   
   IF Sbr_IN_xHeadPos THEN
   	Z300_BufferPlate.rgtPlate[Sbr_IN_dCapIndex].tData.tFlag.tConveyor.xDoneHeadPositioning := 1;
   	IF (Z300_BufferPlate.rgtPlate[Sbr_IN_dCapIndex].tData.dTotalCaps > 1) AND (Z300_BufferPlate.rgtPlate[Sbr_IN_dCapIndex].tTracking.dNextCapIndex > 0) THEN
   		JSR(sbrTrackingPositioningDone,2,Z300_BufferPlate.rgtPlate[Sbr_IN_dCapIndex].tTracking.dNextCapIndex,Sbr_IN_xHeadPos);
   	END_IF;
   ELSE
   	Z300_BufferPlate.rgtPlate[Sbr_IN_dCapIndex].tData.tFlag.tConveyor.xDoneTailPositioning := 1;
   	IF (Z300_BufferPlate.rgtPlate[Sbr_IN_dCapIndex].tData.dTotalCaps > 1) AND (Z300_BufferPlate.rgtPlate[Sbr_IN_dCapIndex].tTracking.dNextCapIndex > 0) THEN
   		JSR(sbrTrackingPositioningDone,2,Z300_BufferPlate.rgtPlate[Sbr_IN_dCapIndex].tTracking.dNextCapIndex,Sbr_IN_xHeadPos);
   	END_IF;
   END_IF;
   
   /*
   Z300_BufferPlate.rgtPlate[Sbr_IN_dCapIndex].tTracking.dPosition_cmm := Sbr_IN_Position - Z300_BufferPlate.rgtPlate[Sbr_IN_dCapIndex].tTracking.dLength_cmm / 2;
   ///////////////// CONVOY SYNCHRONIZATION
   IF (Z300_BufferPlate.rgtPlate[Sbr_IN_dCapIndex].tData.dTotalCaps > 1) AND (Z300_BufferPlate.rgtPlate[Sbr_IN_dCapIndex].tData.dCapIndex = 0) THEN
   	JSR(sbrZ300ConvoySynchronization,1,Sbr_IN_dCapIndex);
   END_IF;
   */
   
END_ROUTINE

ROUTINE sbrTrackingPositioningStart   (* structured text *)
   
   SBR(Sbr_IN_dCapIndex,Sbr_IN_xHeadPos);
   
   IF Sbr_IN_xHeadPos THEN
   	Z300_BufferPlate.rgtPlate[Sbr_IN_dCapIndex].tData.tFlag.tConveyor.xDoneHeadPositioning := 0;
   	IF (Z300_BufferPlate.rgtPlate[Sbr_IN_dCapIndex].tData.dTotalCaps > 1) AND (Z300_BufferPlate.rgtPlate[Sbr_IN_dCapIndex].tTracking.dNextCapIndex > 0) THEN
   		JSR(sbrTrackingPositioningDone,2,Z300_BufferPlate.rgtPlate[Sbr_IN_dCapIndex].tTracking.dNextCapIndex,Sbr_IN_xHeadPos);
   	END_IF;
   ELSE
   	Z300_BufferPlate.rgtPlate[Sbr_IN_dCapIndex].tData.tFlag.tConveyor.xDoneTailPositioning := 0;
   	IF (Z300_BufferPlate.rgtPlate[Sbr_IN_dCapIndex].tData.dTotalCaps > 1) AND (Z300_BufferPlate.rgtPlate[Sbr_IN_dCapIndex].tTracking.dNextCapIndex > 0) THEN
   		JSR(sbrTrackingPositioningDone,2,Z300_BufferPlate.rgtPlate[Sbr_IN_dCapIndex].tTracking.dNextCapIndex,Sbr_IN_xHeadPos);
   	END_IF;
   END_IF;
   
END_ROUTINE

ROUTINE sbrTrackingShift   (* structured text *)
   
   FOR TMP_dIndexCap:=0 TO CONST_tPlant.dMaxNumPlates - 1 DO
   	TMP_xTailFound := 0;
   	TMP_xCenterFound := 0;
   	TMP_OUT_xPlateEndTracking := 0;
   	SIZE(Z300_LineTracking.rgtTrkConv[0],0,TMP_dLineSize);
   
   	//Check Tracking Data Present
   	IF (Z300_BufferPlate.rgtPlate[TMP_dIndexCap].tTracking.dPosition_cmm < Z300_dEndTrackingPosition) AND (Z300_BufferPlate.rgtPlate[TMP_dIndexCap].tTracking.dLength_cmm > 0) THEN
   	    TMP_dStepAdvMotor := Z300_BufferPlate.rgtPlate[TMP_dIndexCap].tTracking.dIndexMotorStepAdv;
   		IF NOT Z300_BufferPlate.rgtPlate[TMP_dIndexCap].tTracking.xNotConsConvTrk THEN
   			IF Z300_BufferPlate.rgtPlate[TMP_dIndexCap].tTracking.dLastConv > 0 THEN
   		        TMP_dLastConv := Z300_BufferPlate.rgtPlate[TMP_dIndexCap].tTracking.dLastConv;
   		        Z300_BufferPlate.rgtPlate[TMP_dIndexCap].tTracking.dLastConv := 0;
   
   		        FOR TMP_dIndexConv := TMP_dLastConv - 1 TO TMP_dLastConv + 1 DO
   		            IF (Z300_BufferPlate.rgtPlate[TMP_dIndexCap].tTracking.dPosition_cmm >= Z300_LineTracking.rgtTrkConv[TMP_dIndexConv].dStartPosition_cmm
   						OR (Z300_BufferPlate.rgtPlate[TMP_dIndexCap].tTracking.dPosition_cmm <= Z300_LineTracking.rgtTrkConv[TMP_dIndexConv].dStartPosition_cmm AND TMP_dIndexConv = 0 ))
   		                   AND Z300_BufferPlate.rgtPlate[TMP_dIndexCap].tTracking.dPosition_cmm <= Z300_LineTracking.rgtTrkConv[TMP_dIndexConv].dEndPosition_cmm THEN
   		                IF NOT Z300_BufferPlate.rgtPlate[TMP_dIndexCap].tTracking.xHoldAdvancement THEN
   							IF Z300_Conveyor_Conf[TMP_dIndexConv].dMotorNumber > 0 THEN
   								TMP_dStepAdvMotor := Z300_BufferPlate.rgtPlate[TMP_dIndexCap].tTracking.dIndexMotorStepAdv;
   							ELSE //One motor presence considerate the plate on the first
   								TMP_dStepAdvMotor := 0;
   							END_IF;
   		                    Z300_BufferPlate.rgtPlate[TMP_dIndexCap].tTracking.dPosition_cmm := Z300_BufferPlate.rgtPlate[TMP_dIndexCap].tTracking.dPosition_cmm + Z300_LineTracking.rgtTrkConv[TMP_dIndexConv].dStepAdv_cmm[TMP_dStepAdvMotor];
   		                END_IF;
   		                Z300_BufferPlate.rgtPlate[TMP_dIndexCap].tTracking.dLastConv := TMP_dIndexConv;
   		                EXIT;
   		            END_IF;
   		        END_FOR;
   
   		     // Global Search
   		     ELSE
   		         FOR TMP_dIndexConv := 0 TO TMP_dLineSize - 1 DO
   		             IF (Z300_BufferPlate.rgtPlate[TMP_dIndexCap].tTracking.dPosition_cmm >= Z300_LineTracking.rgtTrkConv[TMP_dIndexConv].dStartPosition_cmm OR
   		                 (Z300_BufferPlate.rgtPlate[TMP_dIndexCap].tTracking.dPosition_cmm <= Z300_LineTracking.rgtTrkConv[TMP_dIndexConv].dStartPosition_cmm AND TMP_dIndexConv = 0 ))
   		                 AND Z300_BufferPlate.rgtPlate[TMP_dIndexCap].tTracking.dPosition_cmm <= Z300_LineTracking.rgtTrkConv[TMP_dIndexConv].dEndPosition_cmm THEN
   		                IF NOT Z300_BufferPlate.rgtPlate[TMP_dIndexCap].tTracking.xHoldAdvancement THEN
   							IF Z300_Conveyor_Conf[TMP_dIndexConv].dMotorNumber > 0 THEN
   								TMP_dStepAdvMotor := Z300_BufferPlate.rgtPlate[TMP_dIndexCap].tTracking.dIndexMotorStepAdv;
   							ELSE //One motor presence considerate the plate on the first
   								TMP_dStepAdvMotor := 0;
   							END_IF;
   		                    Z300_BufferPlate.rgtPlate[TMP_dIndexCap].tTracking.dPosition_cmm := Z300_BufferPlate.rgtPlate[TMP_dIndexCap].tTracking.dPosition_cmm + Z300_LineTracking.rgtTrkConv[TMP_dIndexConv].dStepAdv_cmm[TMP_dStepAdvMotor];
   		                END_IF;
   		                Z300_BufferPlate.rgtPlate[TMP_dIndexCap].tTracking.dLastConv := TMP_dIndexConv;
   		                EXIT;
   		            END_IF;
   		        END_FOR;
   		    END_IF;
   	    ELSE
   			IF NOT Z300_BufferPlate.rgtPlate[TMP_dIndexCap].tTracking.xHoldAdvancement THEN
               	TMP_dIndexConv := Z300_BufferPlate.rgtPlate[TMP_dIndexCap].tTracking.dIndexConvNotCons;
               	IF Z300_Conveyor_Conf[TMP_dIndexConv].dMotorNumber > 0 THEN
   					TMP_dStepAdvMotor := Z300_BufferPlate.rgtPlate[TMP_dIndexCap].tTracking.dIndexMotorStepAdv;
   				ELSE //One motor presence considerate the plate on the first
   					TMP_dStepAdvMotor := 0;
   				END_IF;
               	Z300_BufferPlate.rgtPlate[TMP_dIndexCap].tTracking.dPosition_cmm := Z300_BufferPlate.rgtPlate[TMP_dIndexCap].tTracking.dPosition_cmm + Z300_LineTracking.rgtTrkConv[TMP_dIndexConv].dStepAdv_cmm[TMP_dStepAdvMotor];
           	END_IF;
           	Z300_BufferPlate.rgtPlate[TMP_dIndexCap].tTracking.dLastConv := TMP_dIndexConv;
   		END_IF;
   
   	    TMP_dLastConvTail := Z300_BufferPlate.rgtPlate[TMP_dIndexCap].tTracking.dLastConvTail;
   	    Z300_BufferPlate.rgtPlate[TMP_dIndexCap].tTracking.dLastConvTail := 0;
   	    TMP_xTailFound := 0;
   	    TMP_xCenterFound := 0;
   	    FOR TMP_dIndexConv := TMP_dLastConvTail TO TMP_dLineSize - 1 DO
   
               TMP_dIndexCapConv := Z300_LineTracking.rgtTrkConv[TMP_dIndexConv].dIndexCaps;// - 1;
   
   			IF TMP_dIndexCapConv < CONST_tPlant.dNumCapsConveyor THEN
   	            TMP_dPosTail_cmm := Z300_BufferPlate.rgtPlate[TMP_dIndexCap].tTracking.dPosition_cmm - (Z300_BufferPlate.rgtPlate[TMP_dIndexCap].tTracking.dLength_cmm / 2);
   	            TMP_dPosHead_cmm := Z300_BufferPlate.rgtPlate[TMP_dIndexCap].tTracking.dPosition_cmm + (Z300_BufferPlate.rgtPlate[TMP_dIndexCap].tTracking.dLength_cmm/ 2);
   	            TMP_dPos_cmm := Z300_BufferPlate.rgtPlate[TMP_dIndexCap].tTracking.dPosition_cmm - (Z300_BufferPlate.rgtPlate[TMP_dIndexCap].tTracking.dLength_cmm / 2);
   
   	            //Tail
   	            IF TMP_dPos_cmm >= Z300_LineTracking.rgtTrkConv[TMP_dIndexConv].dStartPosition_cmm
   					AND TMP_dPos_cmm < Z300_LineTracking.rgtTrkConv[TMP_dIndexConv].dEndPosition_cmm  AND NOT TMP_xTailFound THEN
   	                IF TMP_dPos_cmm >= 0 AND TMP_dPos_cmm < Z300_dEndTrackingPosition THEN
   	                    Z300_LineTracking.rgtTrkConv[TMP_dIndexConv].Cap[TMP_dIndexCapConv].xTail := 1;
   	                    Z300_LineTracking.rgtTrkConv[TMP_dIndexConv].Cap[TMP_dIndexCapConv].xPresence := 1;
   	                    Z300_LineTracking.rgtTrkConv[TMP_dIndexConv].Cap[TMP_dIndexCapConv].dTailPos_cmm := TMP_dPos_cmm;
   	                    Z300_LineTracking.rgtTrkConv[TMP_dIndexConv].Cap[TMP_dIndexCapConv].dTailPosConv_cmm := TMP_dPos_cmm - Z300_LineTracking.rgtTrkConv[TMP_dIndexConv].dStartPosition_cmm;
   	                    Z300_LineTracking.rgtTrkConv[TMP_dIndexConv].Cap[TMP_dIndexCapConv].dPointer := TMP_dIndexCap;
   	                    Z300_LineTracking.rgtTrkConv[TMP_dIndexConv].Cap[TMP_dIndexCapConv].dPresenceHead_cmm := TMP_dPosHead_cmm;
   	                    Z300_LineTracking.rgtTrkConv[TMP_dIndexConv].Cap[TMP_dIndexCapConv].dPresenceTail_cmm := TMP_dPosTail_cmm;
   	                    Z300_BufferPlate.rgtPlate[TMP_dIndexCap].tTracking.dIndexConvTail := TMP_dIndexConv;
   	                    TMP_xTailFound := 1;
   	                    Z300_BufferPlate.rgtPlate[TMP_dIndexCap].tTracking.dLastConvTail := TMP_dIndexConv;
   	                    Z300_BufferPlate.rgtPlate[TMP_dIndexCap].tTracking.dIndexCapInConvTail := TMP_dIndexCap;
   	                    Z300_BufferPlate.rgtPlate[TMP_dIndexCap].tTracking.dPositionTail_cmm := TMP_dPos_cmm;
   	                END_IF;
   	            END_IF;
   
   	            // Center Position
   	            TMP_dPosTail_cmm := Z300_BufferPlate.rgtPlate[TMP_dIndexCap].tTracking.dPosition_cmm - (Z300_BufferPlate.rgtPlate[TMP_dIndexCap].tTracking.dLength_cmm / 2);
   	            TMP_dPosHead_cmm := Z300_BufferPlate.rgtPlate[TMP_dIndexCap].tTracking.dPosition_cmm + (Z300_BufferPlate.rgtPlate[TMP_dIndexCap].tTracking.dLength_cmm / 2);
   	            TMP_dPos_cmm := Z300_BufferPlate.rgtPlate[TMP_dIndexCap].tTracking.dPosition_cmm;
   	            IF TMP_dPos_cmm >= Z300_LineTracking.rgtTrkConv[TMP_dIndexConv].dStartPosition_cmm
   					AND TMP_dPos_cmm < Z300_LineTracking.rgtTrkConv[TMP_dIndexConv].dEndPosition_cmm AND NOT TMP_xCenterFound THEN
   	                IF TMP_dPos_cmm >= Z300_dStartTrackingPosition AND TMP_dPos_cmm < Z300_dEndTrackingPosition THEN
   	                    Z300_LineTracking.rgtTrkConv[TMP_dIndexConv].Cap[TMP_dIndexCapConv].xCenter := 1;
   	                    Z300_LineTracking.rgtTrkConv[TMP_dIndexConv].Cap[TMP_dIndexCapConv].xPresence := 1;
   	                    Z300_LineTracking.rgtTrkConv[TMP_dIndexConv].Cap[TMP_dIndexCapConv].dCenterPos_cmm := TMP_dPos_cmm;
   	                    Z300_LineTracking.rgtTrkConv[TMP_dIndexConv].Cap[TMP_dIndexCapConv].dCenterPosConv_cmm := TMP_dPos_cmm - Z300_LineTracking.rgtTrkConv[TMP_dIndexConv].dStartPosition_cmm;
   	                    Z300_LineTracking.rgtTrkConv[TMP_dIndexConv].Cap[TMP_dIndexCapConv].dPointer := TMP_dIndexCap;
   	                    Z300_LineTracking.rgtTrkConv[TMP_dIndexConv].Cap[TMP_dIndexCapConv].dPresenceHead_cmm := TMP_dPosHead_cmm;
   	                    Z300_LineTracking.rgtTrkConv[TMP_dIndexConv].Cap[TMP_dIndexCapConv].dPresenceTail_cmm := TMP_dPosTail_cmm;
   	                    TMP_xCenterFound := 1;
   	                END_IF;
   	            END_IF;
   
   	            //Plate Presence
   	            TMP_dPosTail_cmm := Z300_BufferPlate.rgtPlate[TMP_dIndexCap].tTracking.dPosition_cmm - (Z300_BufferPlate.rgtPlate[TMP_dIndexCap].tTracking.dLength_cmm / 2);
   	            TMP_dPosHead_cmm := Z300_BufferPlate.rgtPlate[TMP_dIndexCap].tTracking.dPosition_cmm + (Z300_BufferPlate.rgtPlate[TMP_dIndexCap].tTracking.dLength_cmm / 2);
   	            IF TMP_dPosTail_cmm <= Z300_LineTracking.rgtTrkConv[TMP_dIndexConv].dStartPosition_cmm
   					AND TMP_dPosHead_cmm >= Z300_LineTracking.rgtTrkConv[TMP_dIndexConv].dEndPosition_cmm  THEN
   	                IF TMP_dPos_cmm >= Z300_dStartTrackingPosition AND TMP_dPos_cmm < Z300_dEndTrackingPosition THEN
   	                    Z300_LineTracking.rgtTrkConv[TMP_dIndexConv].Cap[TMP_dIndexCapConv].xPresence := 1;
   	                    Z300_LineTracking.rgtTrkConv[TMP_dIndexConv].Cap[TMP_dIndexCapConv].dCenterPos_cmm := TMP_dPos_cmm;
   	                    Z300_LineTracking.rgtTrkConv[TMP_dIndexConv].Cap[TMP_dIndexCapConv].dPresenceHead_cmm := TMP_dPosHead_cmm;
   	                    Z300_LineTracking.rgtTrkConv[TMP_dIndexConv].Cap[TMP_dIndexCapConv].dPresenceTail_cmm := TMP_dPosTail_cmm;
   	                    Z300_LineTracking.rgtTrkConv[TMP_dIndexConv].Cap[TMP_dIndexCapConv].dCenterPosConv_cmm := TMP_dPos_cmm - Z300_LineTracking.rgtTrkConv[TMP_dIndexConv].dStartPosition_cmm;
   	                    Z300_LineTracking.rgtTrkConv[TMP_dIndexConv].Cap[TMP_dIndexCapConv].dPointer := TMP_dIndexCap;
   	                    TMP_xPlateFound := 1;
   	                END_IF;
   	            END_IF;
   
   	            // Head Position
   	            TMP_dPosTail_cmm := Z300_BufferPlate.rgtPlate[TMP_dIndexCap].tTracking.dPosition_cmm - (Z300_BufferPlate.rgtPlate[TMP_dIndexCap].tTracking.dLength_cmm / 2);
   	            TMP_dPosHead_cmm := Z300_BufferPlate.rgtPlate[TMP_dIndexCap].tTracking.dPosition_cmm + (Z300_BufferPlate.rgtPlate[TMP_dIndexCap].tTracking.dLength_cmm / 2);
   	            TMP_dPos_cmm := Z300_BufferPlate.rgtPlate[TMP_dIndexCap].tTracking.dPosition_cmm + (Z300_BufferPlate.rgtPlate[TMP_dIndexCap].tTracking.dLength_cmm / 2);
   	            IF (TMP_dPos_cmm >= Z300_LineTracking.rgtTrkConv[TMP_dIndexConv].dStartPosition_cmm)
   					AND (TMP_dPos_cmm < Z300_LineTracking.rgtTrkConv[TMP_dIndexConv].dEndPosition_cmm) AND TMP_xCenterFound THEN
   	                IF TMP_dPos_cmm >= Z300_dStartTrackingPosition AND TMP_dPos_cmm < Z300_dEndTrackingPosition THEN
   	                    Z300_LineTracking.rgtTrkConv[TMP_dIndexConv].Cap[TMP_dIndexCapConv].xHead := 1;
   	                    Z300_LineTracking.rgtTrkConv[TMP_dIndexConv].Cap[TMP_dIndexCapConv].xPresence := 1;
   	                    Z300_LineTracking.rgtTrkConv[TMP_dIndexConv].Cap[TMP_dIndexCapConv].dHeadPos_cmm := TMP_dPos_cmm;
   	                    Z300_LineTracking.rgtTrkConv[TMP_dIndexConv].Cap[TMP_dIndexCapConv].dHeadPosConv_cmm := TMP_dPos_cmm - Z300_LineTracking.rgtTrkConv[TMP_dIndexConv].dStartPosition_cmm;
   	                    Z300_LineTracking.rgtTrkConv[TMP_dIndexConv].Cap[TMP_dIndexCapConv].dPointer := TMP_dIndexCap;
   	                    Z300_LineTracking.rgtTrkConv[TMP_dIndexConv].Cap[TMP_dIndexCapConv].dPresenceHead_cmm := TMP_dPosHead_cmm;
   	                    Z300_LineTracking.rgtTrkConv[TMP_dIndexConv].Cap[TMP_dIndexCapConv].dPresenceTail_cmm := TMP_dPosTail_cmm;
   	                    //Increment Index Single Caps in the conveyor
   	                    Z300_LineTracking.rgtTrkConv[TMP_dIndexConv].dIndexCaps := Z300_LineTracking.rgtTrkConv[TMP_dIndexConv].dIndexCaps + 1;
   	                    IF Z300_LineTracking.rgtTrkConv[TMP_dIndexConv].dIndexCaps >= CONST_tPlant.dNumCapsConveyor THEN
   	                        Z300_LineTracking.rgtTrkConv[TMP_dIndexConv].dIndexCaps := CONST_tPlant.dNumCapsConveyor - 1;
   	                    END_IF;
   	                    Z300_BufferPlate.rgtPlate[TMP_dIndexCap].tTracking.dIndexConvHead := TMP_dIndexConv;
   	                    Z300_BufferPlate.rgtPlate[TMP_dIndexCap].tTracking.dIndexCapInConvHead := TMP_dIndexCap;
   	                    Z300_BufferPlate.rgtPlate[TMP_dIndexCap].tTracking.dPositionHead_cmm := TMP_dPos_cmm;
   	                    EXIT;
   	                END_IF;
   	            END_IF;
   
   			END_IF;
   
               IF  TMP_xTailFound OR TMP_xCenterFound OR TMP_xPlateFound THEN
                   //Increment Index Single Caps in the conveyor
                   Z300_LineTracking.rgtTrkConv[TMP_dIndexConv].dIndexCaps := Z300_LineTracking.rgtTrkConv[TMP_dIndexConv].dIndexCaps + 1;
                   IF Z300_LineTracking.rgtTrkConv[TMP_dIndexConv].dIndexCaps >= CONST_tPlant.dNumCapsConveyor THEN
                       Z300_LineTracking.rgtTrkConv[TMP_dIndexConv].dIndexCaps := CONST_tPlant.dNumCapsConveyor - 1;
                   END_IF;
               END_IF;
           END_FOR;
       ELSE
   		//plate not more in tracking area
   		TMP_OUT_xPlateEndTracking := Z300_BufferPlate.rgtPlate[TMP_dIndexCap].tTracking.dPosition_cmm >= Z300_dEndTrackingPosition;
   	END_IF;
   
       //write the Output
       Z300_BufferPlate.rgtPlate[TMP_dIndexCap].tTracking.dPosition_cmm := Z300_BufferPlate.rgtPlate[TMP_dIndexCap].tTracking.dPosition_cmm;
   
   	//if plate at end of tracking delete from tracking
   	IF TMP_OUT_xPlateEndTracking THEN
   		COP(AUX_tBufferPlate_NULL,Z300_BufferPlate.rgtPlate[TMP_dIndexCap],1);
   	END_IF;
   END_FOR;
   
END_ROUTINE

ROUTINE sbrTrimWheelTrPositionOppOpSide   (* ladder *)
   0: NOP();
   1: [XIC(M30xTrimWheel[TMP_dIndex].OS_xStartPositioningOppOpSide) ,XIC(M30xTrimWheel[TMP_dIndex].OS_xReqUpdateTargetTranslationOppOpSide) ]ADD(M30xTrimWheel[TMP_dIndex].AUX_dReqTargetPosTranslation_cmm[1],M30xTrimWheel[TMP_dIndex].AUX_dOffsetSingle_cmm[1],M30xTrimWheel[TMP_dIndex].AUX_dFinalTarget_cmm[1]);
   2: GP_PosWindow(GP_PosWindow,M30xTrimWheel[TMP_dIndex].AUX_dFinalTarget_cmm[1],M30xTrimWheel[TMP_dIndex].AUX_dActTransPosition_cmm[1],M30xTrimWheel[TMP_dIndex].CONF_dTolerance_cmm[1],0,M30xTrimWheel[TMP_dIndex].ST_xInPositionOppOpSide);
   3: GP_PosWindow(GP_PosWindow,M30xTrimWheel[TMP_dIndex].AUX_dFinalTarget_cmm[1],M30xTrimWheel[TMP_dIndex].AUX_dActTransPosition_cmm[1],M30xTrimWheel[TMP_dIndex].CONF_dStopCamPos_cmm[1],0,M30xTrimWheel[TMP_dIndex].ST_xInStopCamPositionOppOpSide);
   4: GP_PosWindow(GP_PosWindow,M30xTrimWheel_HMW[TMP_dIndex].rgdPositionManCmd_cmm[1],M30xTrimWheel[TMP_dIndex].AUX_dActTransPosition_cmm[1],M30xTrimWheel[TMP_dIndex].CONF_dSlowDownPos_cmm[1],0,M30xTrimWheel[TMP_dIndex].ST_xInSlowDownManualPosOppOpSide);
   5: GP_PosWindow(GP_PosWindow,M30xTrimWheel_HMW[TMP_dIndex].rgdPositionManCmd_cmm[1],M30xTrimWheel[TMP_dIndex].AUX_dActTransPosition_cmm[1],M30xTrimWheel[TMP_dIndex].CONF_dStopCamPos_cmm[1],0,M30xTrimWheel[TMP_dIndex].ST_xInStopCamManualPositionOppOpSide);
   6: XIC(M30xTrimWheel_HMW[TMP_dIndex].rgxMan.x12)MOV(M30xTrimWheel[TMP_dIndex].CONF_dTrimWheelMaxRange_cmm[1],TMP_dManualTargetPos);
   7: XIC(M30xTrimWheel_HMW[TMP_dIndex].rgxMan.x13)MOV(M30xTrimWheel[TMP_dIndex].CONF_dTrimWheelMinRange_cmm[1],TMP_dManualTargetPos);
   8: GP_PosWindow(GP_PosWindow,TMP_dManualTargetPos,M30xTrimWheel[TMP_dIndex].AUX_dActTransPosition_cmm[1],M30xTrimWheel[TMP_dIndex].CONF_dSlowDownPos_cmm[1],0,M30xTrimWheel[TMP_dIndex].ST_xInSlowDownManualOppOpSide);
   9: GP_PosWindow(GP_PosWindow,TMP_dManualTargetPos,M30xTrimWheel[TMP_dIndex].AUX_dActTransPosition_cmm[1],M30xTrimWheel[TMP_dIndex].CONF_dStopCamPos_cmm[1],0,M30xTrimWheel[TMP_dIndex].ST_xInStopCamManualOppOpSide);
END_ROUTINE

ROUTINE sbrTrimWheelTrPositionOpSide   (* ladder *)
   0: NOP();
   1: [XIC(M30xTrimWheel[TMP_dIndex].OS_xStartPositioningOpSide) ,XIC(M30xTrimWheel[TMP_dIndex].OS_xReqUpdateTargetTranslationOpSide) ]ADD(M30xTrimWheel[TMP_dIndex].AUX_dReqTargetPosTranslation_cmm[0],M30xTrimWheel[TMP_dIndex].AUX_dOffsetSingle_cmm[0],M30xTrimWheel[TMP_dIndex].AUX_dFinalTarget_cmm[0]);
   2: GP_PosWindow(GP_PosWindow,M30xTrimWheel[TMP_dIndex].AUX_dFinalTarget_cmm[0],M30xTrimWheel[TMP_dIndex].AUX_dActTransPosition_cmm[0],M30xTrimWheel[TMP_dIndex].CONF_dTolerance_cmm[0],0,M30xTrimWheel[TMP_dIndex].ST_xInPositionOpSide);
   3: GP_PosWindow(GP_PosWindow,M30xTrimWheel[TMP_dIndex].AUX_dFinalTarget_cmm[0],M30xTrimWheel[TMP_dIndex].AUX_dActTransPosition_cmm[0],M30xTrimWheel[TMP_dIndex].CONF_dStopCamPos_cmm[0],0,M30xTrimWheel[TMP_dIndex].ST_xInStopCamPositionOpSide);
   4: GP_PosWindow(GP_PosWindow,M30xTrimWheel_HMW[TMP_dIndex].rgdPositionManCmd_cmm[0],M30xTrimWheel[TMP_dIndex].AUX_dActTransPosition_cmm[0],M30xTrimWheel[TMP_dIndex].CONF_dSlowDownPos_cmm[0],0,M30xTrimWheel[TMP_dIndex].ST_xInSlowDownManualPosOpSide);
   5: GP_PosWindow(GP_PosWindow,M30xTrimWheel_HMW[TMP_dIndex].rgdPositionManCmd_cmm[0],M30xTrimWheel[TMP_dIndex].AUX_dActTransPosition_cmm[0],M30xTrimWheel[TMP_dIndex].CONF_dStopCamPos_cmm[0],0,M30xTrimWheel[TMP_dIndex].ST_xInStopCamManualPositionOpSide);
   6: XIC(M30xTrimWheel_HMW[TMP_dIndex].rgxMan.x2)MOV(M30xTrimWheel[TMP_dIndex].CONF_dTrimWheelMaxRange_cmm[0],TMP_dManualTargetPos);
   7: XIC(M30xTrimWheel_HMW[TMP_dIndex].rgxMan.x3)MOV(M30xTrimWheel[TMP_dIndex].CONF_dTrimWheelMinRange_cmm[0],TMP_dManualTargetPos);
   8: GP_PosWindow(GP_PosWindow,TMP_dManualTargetPos,M30xTrimWheel[TMP_dIndex].AUX_dActTransPosition_cmm[0],M30xTrimWheel[TMP_dIndex].CONF_dSlowDownPos_cmm[0],0,M30xTrimWheel[TMP_dIndex].ST_xInSlowDownManualOpSide);
   9: GP_PosWindow(GP_PosWindow,TMP_dManualTargetPos,M30xTrimWheel[TMP_dIndex].AUX_dActTransPosition_cmm[0],M30xTrimWheel[TMP_dIndex].CONF_dStopCamPos_cmm[0],0,M30xTrimWheel[TMP_dIndex].ST_xInStopCamManualOpSide);
END_ROUTINE

ROUTINE sbrUpdateTrackingConvoyPosition   (* structured text *)
   SBR(Sbr_IN_dIndexHead,Sbr_IN_Position);
   
   Z300_BufferPlate.rgtPlate[Sbr_IN_dIndexHead].tTracking.dPosition_cmm := Sbr_IN_Position - Z300_BufferPlate.rgtPlate[Sbr_IN_dIndexHead].tTracking.dLength_cmm / 2;
   ///////////////// CONVOY SYNCHRONIZATION
   IF (Z300_BufferPlate.rgtPlate[Sbr_IN_dIndexHead].tData.dTotalCaps > 1) AND (Z300_BufferPlate.rgtPlate[Sbr_IN_dIndexHead].tData.dCapIndex = 0) THEN
   //Search for single caps within the same convoy
   	// Synchronize convoy
   	JSR(sbrZ300ConvoySynchronization,1,Sbr_IN_dIndexHead);
   END_IF;
   
END_ROUTINE

ROUTINE sbrZ300ConvoySynchronization   (* structured text *)
   /*
   //Initialize
   TMP_dPnt1 := Z300_Photocell[TMP_dIndex].tSearchPlate.rgdHeadPointer[0];
   TMP_dPnt2 := Z300_Photocell[TMP_dIndex].tSearchPlate.rgdHeadPointer[1];
   TMP_dPnt3 := Z300_Photocell[TMP_dIndex].tSearchPlate.rgdHeadPointer[2];
   TMP_dPnt4 := Z300_Photocell[TMP_dIndex].tSearchPlate.rgdHeadPointer[3];
   //If convoy in progress synchronize second cap
   IF (Z300_Photocell[TMP_dIndex].tSearchPlate.rgxHead > 1) AND (Z300_BufferPlate.rgtPlate[TMP_dPnt1].tData.dTotalCaps > 1) AND (Z300_BufferPlate.rgtPlate[TMP_dPnt1].tData.rgtCap[0].dIndex = 0)
   AND (Z300_BufferPlate.rgtPlate[TMP_dPnt2].tData.dTotalCaps > 1) AND (Z300_BufferPlate.rgtPlate[TMP_dPnt2].tData.rgtCap[0].dIndex = 1) THEN
   	//Synchronyze also second cap
   	Z300_BufferPlate.rgtPlate[TMP_dPnt2].tTracking.dPosition_cmm := Z300_BufferPlate.rgtPlate[TMP_dPnt1].tTracking.dPosition_cmm
   	- (Z300_BufferPlate.rgtPlate[TMP_dPnt1].tTracking.dLength_cmm / 2)
   	- Z300_BufferPlate.rgtPlate[TMP_dPnt1].tData.dGapCaps_cmm
   	- (Z300_BufferPlate.rgtPlate[TMP_dPnt2].tTracking.dLength_cmm / 2);
   END_IF;
   //If convoy in progress synchronize third cap
   IF (Z300_Photocell[TMP_dIndex].tSearchPlate.rgxHead > 2) AND (Z300_BufferPlate.rgtPlate[TMP_dPnt2].tData.dTotalCaps > 2) AND (Z300_BufferPlate.rgtPlate[TMP_dPnt2].tData.rgtCap[0].dIndex = 1)
   AND (Z300_BufferPlate.rgtPlate[TMP_dPnt3].tData.dTotalCaps > 2) AND (Z300_BufferPlate.rgtPlate[TMP_dPnt3].tData.rgtCap[0].dIndex = 2) THEN
   	//Synchronyze also third cap
   	Z300_BufferPlate.rgtPlate[TMP_dPnt3].tTracking.dPosition_cmm := Z300_BufferPlate.rgtPlate[TMP_dPnt2].tTracking.dPosition_cmm
   	- (Z300_BufferPlate.rgtPlate[TMP_dPnt2].tTracking.dLength_cmm / 2)
   	- Z300_BufferPlate.rgtPlate[TMP_dPnt2].tData.dGapCaps_cmm
   	- (Z300_BufferPlate.rgtPlate[TMP_dPnt3].tTracking.dLength_cmm / 2);
   END_IF;
   //If convoy in progress synchronize fourth cap
   IF (Z300_Photocell[TMP_dIndex].tSearchPlate.rgxHead > 3) AND (Z300_BufferPlate.rgtPlate[TMP_dPnt3].tData.dTotalCaps > 3) AND (Z300_BufferPlate.rgtPlate[TMP_dPnt3].tData.rgtCap[0].dIndex = 2)
   AND (Z300_BufferPlate.rgtPlate[TMP_dPnt4].tData.dTotalCaps > 3) AND (Z300_BufferPlate.rgtPlate[TMP_dPnt4].tData.rgtCap[0].dIndex = 3) THEN
   	//Synchronyze also fourth cap
   	Z300_BufferPlate.rgtPlate[TMP_dPnt4].tTracking.dPosition_cmm := Z300_BufferPlate.rgtPlate[TMP_dPnt3].tTracking.dPosition_cmm
   	- (Z300_BufferPlate.rgtPlate[TMP_dPnt3].tTracking.dLength_cmm / 2)
   	- Z300_BufferPlate.rgtPlate[TMP_dPnt3].tData.dGapCaps_cmm
   	- (Z300_BufferPlate.rgtPlate[TMP_dPnt4].tTracking.dLength_cmm / 2);
   END_IF;
   */
   
   SBR(Sbr_IN_dCapIndex);
   
   TMP_dNextCap := Z300_BufferPlate.rgtPlate[Sbr_IN_dCapIndex].tTracking.dNextCapIndex;
   IF TMP_dNextCap > 0 THEN
   	Z300_BufferPlate.rgtPlate[TMP_dNextCap].tTracking.dPosition_cmm := Z300_BufferPlate.rgtPlate[Sbr_IN_dCapIndex].tTracking.dPosition_cmm - Z300_BufferPlate.rgtPlate[Sbr_IN_dCapIndex].tTracking.dLength_cmm / 2
   	- Z300_BufferPlate.rgtPlate[Sbr_IN_dCapIndex].tData.dGapCaps_cmm - Z300_BufferPlate.rgtPlate[TMP_dNextCap].tTracking.dLength_cmm / 2;
   	JSR(sbrZ300ConvoySynchronization,1,TMP_dNextCap);
   END_IF;
   
END_ROUTINE

ROUTINE ScadaPlate_Logic   (* structured text *)
   
   TMP_xLastModalityLoadBwd := 0;
   TMP_xLastModalityUnloadBwd := 0;
   TMP_xYWithBarycenter := 1;
   TMP_xYInversionLite := 1;
   
   TMP_dCulletMask := CONST_rgdDestMask[24];
   FOR TMP_dIndexPlate := 0 TO CONST_tPlant.dMaxNumPlates - 1 DO
   	//Write data
   	//Calculate Head Position
   	TMP_dHeadPosition_mm := Z300_BufferPlate.rgtPlate[TMP_dIndexPlate].tTracking.dPositionHead_cmm / 100;
   	TMP_dConveyorLength := Z300_dEndTrackingPosition/ 100;
   	TMP_dWidth_mm := Z300_Conveyor_Conf[0].dWidthConveyor_cmm / 100;
   
   	//Init counter cap (always only one cap on line tracking)
   	TMP_dCap := 0;
   
   	//Init counter lite
   	TMP_dLite := 0;
   
   	FOR TMP_dLite := 0 TO CONST_tPlant.dNumLitesMaxCap - 1 DO
   	    IF Z300_BufferPlate.rgtPlate[TMP_dIndexPlate].tData.rgtCap[TMP_dCap].rgtLite[TMP_dLite].dID <> 0 AND NOT Z300_BufferPlate.rgtPlate[TMP_dIndexPlate].tTracking.xNotShownInScada THEN
   	        TMP_dLiteInv := CONST_tPlant.dNumLitesMaxCap - 1 - TMP_dLite;
   
   	        //Plate
   	        Z300_Scada_Continuous.rgtPlate[TMP_dIndexPlate].rgtCap[TMP_dCap].rgtLite[TMP_dLite].dPlateId := Z300_BufferPlate.rgtPlate[TMP_dIndexPlate].tData.rgtCap[TMP_dCap].rgtLite[TMP_dLite].dID;
   	        //Production ID
   	        Z300_Scada_Continuous.rgtPlate[TMP_dIndexPlate].rgtCap[TMP_dCap].rgtLite[TMP_dLite].dProductionID := Z300_BufferPlate.rgtPlate[TMP_dIndexPlate].tData.rgtCap[TMP_dCap].rgtLite[TMP_dLite].dProductionID;
   	        //Plate lenght
   	        Z300_Scada_Continuous.rgtPlate[TMP_dIndexPlate].rgtCap[TMP_dCap].rgtLite[TMP_dLite].dPlateLength_mm := Z300_BufferPlate.rgtPlate[TMP_dIndexPlate].tData.rgtCap[TMP_dCap].dLength_cmm / 100;
   	        //Plate widht
   	        Z300_Scada_Continuous.rgtPlate[TMP_dIndexPlate].rgtCap[TMP_dCap].rgtLite[TMP_dLite].dPlateWidth_mm := Z300_BufferPlate.rgtPlate[TMP_dIndexPlate].tData.rgtCap[TMP_dCap].rgtLite[TMP_dLite].dWidth_cmm / 100;
   
   	        //Init the value of Destination/Source/Alternative/SecondDestination
   	        TMP_xPresenceDestination := 0;
   	        TMP_xPresenceAlternative := 0;
   	        //TMP_xPresenceSource := 0;
   	        TMP_xPresenceSecondDestination := 0;
   
   	        //Destination
   	        FOR TMP_dCountDest := 0 TO 31 DO
   	            //Main Destination
   	            IF Z300_BufferPlate.rgtPlate[TMP_dIndexPlate].tData.rgtCap[TMP_dCap].rgtLite[TMP_dLite].tDestination.rgxMain.[TMP_dCountDest] THEN
   	                Z300_Scada_Continuous.rgtPlate[TMP_dIndexPlate].rgtCap[TMP_dCap].rgtLite[TMP_dLite].dDestination := TMP_dCountDest + 1;
   	                TMP_xPresenceDestination := 1;
   	            END_IF;
   	            ////Source
   				//IF INO_tPlate.tData.rgtCap[TMP_dCap].rgtLite[TMP_dLite].
   	            //IF INO_tPlate.tData.rgtCap[TMP_dCap].rgtLite[TMP_dLite].tSource.rgxOrigin.[TMP_dCountDest] THEN
   	            //    INO_tScada_Continuous.rgtPlate[IN_dIndexPlate].rgtCap[TMP_dCap].rgtLite[TMP_dLite].dSource := TMP_dCountDest + 1;
   	            //    TMP_xPresenceSource := 1;
   	            //END_IF;
   	            //Alternative Destination
   	            IF Z300_BufferPlate.rgtPlate[TMP_dIndexPlate].tData.rgtCap[TMP_dCap].rgtLite[TMP_dLite].tDestination.rgxAlternative.[TMP_dCountDest] THEN
   	                Z300_Scada_Continuous.rgtPlate[TMP_dIndexPlate].rgtCap[TMP_dCap].rgtLite[TMP_dLite].dAlternative := TMP_dCountDest + 1;
   	                TMP_xPresenceAlternative := 1;
   	            END_IF;
   	            //Second Destination
   	            IF Z300_BufferPlate.rgtPlate[TMP_dIndexPlate].tData.rgtCap[TMP_dCap].rgtLite[TMP_dLite].tDestination.rgxAlternative.[TMP_dCountDest] THEN
   	                Z300_Scada_Continuous.rgtPlate[TMP_dIndexPlate].rgtCap[TMP_dCap].rgtLite[TMP_dLite].dSecondDestination := TMP_dCountDest + 1;
   	                TMP_xPresenceSecondDestination := 1;
   	            END_IF;
   	        END_FOR;
   			//IF Z300_BufferPlate.rgtPlate[TMP_dIndexPlate].tData.rgtCap[TMP_dCap].rgtLite[TMP_dLite].tDestination.rgxMain = CONST_rgdDestMask[24] THEN
   	        //    Z300_Scada_Continuous.rgtPlate[TMP_dIndexPlate].rgtCap[TMP_dCap].rgtLite[TMP_dLite].dDestination := CONST_rgdDestMask[24];
   	        //END_IF;
   	        IF NOT TMP_xPresenceDestination THEN
   	            Z300_Scada_Continuous.rgtPlate[TMP_dIndexPlate].rgtCap[TMP_dCap].rgtLite[TMP_dLite].dDestination := 0;
   	        END_IF;
   	        IF NOT TMP_xPresenceAlternative THEN
   	            Z300_Scada_Continuous.rgtPlate[TMP_dIndexPlate].rgtCap[TMP_dCap].rgtLite[TMP_dLite].dAlternative := 0;
   	        END_IF;
   	        IF NOT TMP_xPresenceSecondDestination THEN
   	            Z300_Scada_Continuous.rgtPlate[TMP_dIndexPlate].rgtCap[TMP_dCap].rgtLite[TMP_dLite].dSecondDestination := 0;
   	        END_IF;
   	        //IF NOT TMP_xPresenceSource THEN
   	            Z300_Scada_Continuous.rgtPlate[TMP_dIndexPlate].rgtCap[TMP_dCap].rgtLite[TMP_dLite].dSource := 0;
   	        //END_IF;
   
   	        ////Set origin to 0 in case of destination is <> 0
   	        //IF INO_tScada_Continuous.rgtPlate[IN_dIndexPlate].rgtCap[TMP_dCap].rgtLite[TMP_dLite].dDestination <> 0 THEN
   	        //    INO_tScada_Continuous.rgtPlate[IN_dIndexPlate].rgtCap[TMP_dCap].rgtLite[TMP_dLite].dSource := 0;
   	        //END_IF;
   
   	        //Position x (Forward)
   	        IF NOT TMP_xLastModalityLoadBwd AND NOT TMP_xLastModalityUnloadBwd THEN
   	            //Tail
   	            Z300_Scada_Continuous.rgtPlate[TMP_dIndexPlate].rgtCap[TMP_dCap].rgtLite[TMP_dLite].dTail_PosX_mm := TMP_dHeadPosition_mm - (Z300_BufferPlate.rgtPlate[TMP_dIndexPlate].tData.rgtCap[TMP_dCap].dLength_cmm / 100);
   
   	            //Head
   	            Z300_Scada_Continuous.rgtPlate[TMP_dIndexPlate].rgtCap[TMP_dCap].rgtLite[TMP_dLite].dHead_PosX_mm := TMP_dHeadPosition_mm;
   	        END_IF;
   
   	        //Position x (Backward)
   	        //Head
   
   	        IF TMP_xLastModalityLoadBwd OR TMP_xLastModalityUnloadBwd THEN
   	            //  Head
   	            Z300_Scada_Continuous.rgtPlate[TMP_dIndexPlate].rgtCap[TMP_dCap].rgtLite[TMP_dLite].dHead_PosX_mm := TMP_dConveyorLength - TMP_dHeadPosition_mm + (Z300_BufferPlate.rgtPlate[TMP_dIndexPlate].tData.dLength_cmm / 100);
   
   	            //  Tail
   	            Z300_Scada_Continuous.rgtPlate[TMP_dIndexPlate].rgtCap[TMP_dCap].rgtLite[TMP_dLite].dTail_PosX_mm :=
   	            Z300_Scada_Continuous.rgtPlate[TMP_dIndexPlate].rgtCap[TMP_dCap].rgtLite[TMP_dLite].dHead_PosX_mm - (Z300_BufferPlate.rgtPlate[TMP_dIndexPlate].tData.rgtCap[TMP_dCap].dLength_cmm / 100);
   	        END_IF;
   
   	        //Position Y
   
   	        //Barycenter not used, without inversion (IN FC)
   	        IF NOT TMP_xYWithBarycenter AND NOT TMP_xYInversionLite THEN
   	            IF TMP_dLite < 1 THEN
   	                Z300_Scada_Continuous.rgtPlate[TMP_dIndexPlate].rgtCap[TMP_dCap].rgtLite[TMP_dLite].dPositionY_mm :=
   	                ((TMP_dWidth_mm / 2) - (Z300_BufferPlate.rgtPlate[TMP_dIndexPlate].tData.rgtCap[TMP_dCap].dWidth_cmm / 100) / 2);
   	            ELSE
   	                Z300_Scada_Continuous.rgtPlate[TMP_dIndexPlate].rgtCap[TMP_dCap].rgtLite[TMP_dLite].dPositionY_mm := Z300_Scada_Continuous.rgtPlate[TMP_dIndexPlate].rgtCap[TMP_dCap].rgtLite[TMP_dLite - 1].dPositionY_mm
   	                + (Z300_BufferPlate.rgtPlate[TMP_dIndexPlate].tData.rgtCap[TMP_dCap].rgtLite[TMP_dLite - 1].dWidth_cmm / 100) +
   	                (Z300_BufferPlate.rgtPlate[TMP_dIndexPlate].tData.rgtCap[TMP_dCap].dGap_cmm / 100);
   	            END_IF;
   	        END_IF;
   
   	        //Barycenter not used, with inversion (IN FC)
   	        IF NOT TMP_xYWithBarycenter AND TMP_xYInversionLite THEN
   	            IF TMP_dLite < 1 THEN
   	                Z300_Scada_Continuous.rgtPlate[TMP_dIndexPlate].rgtCap[TMP_dCap].rgtLite[TMP_dLite].dPositionY_mm :=
   	                (TMP_dWidth_mm / 2) + ((Z300_BufferPlate.rgtPlate[TMP_dIndexPlate].tData.rgtCap[TMP_dCap].dWidth_cmm / 100) / 2) -
   	                (Z300_BufferPlate.rgtPlate[TMP_dIndexPlate].tData.rgtCap[TMP_dCap].rgtLite[TMP_dLite].dWidth_cmm / 100);
   
   	            ELSE
   	                Z300_Scada_Continuous.rgtPlate[TMP_dIndexPlate].rgtCap[TMP_dCap].rgtLite[TMP_dLite].dPositionY_mm := Z300_Scada_Continuous.rgtPlate[TMP_dIndexPlate].rgtCap[TMP_dCap].rgtLite[TMP_dLite - 1].dPositionY_mm
   	                - (Z300_BufferPlate.rgtPlate[TMP_dIndexPlate].tData.rgtCap[TMP_dCap].rgtLite[TMP_dLite].dWidth_cmm / 100) -
   	                (Z300_BufferPlate.rgtPlate[TMP_dIndexPlate].tData.rgtCap[TMP_dCap].dGap_cmm / 100);
   	            END_IF;
   	        END_IF;
   
   	        //Barycenter used, without inversion (IN FC)
   
   	        IF TMP_xYWithBarycenter AND NOT TMP_xYInversionLite THEN
   	            Z300_Scada_Continuous.rgtPlate[TMP_dIndexPlate].rgtCap[TMP_dCap].rgtLite[TMP_dLite].dPositionY_mm :=
   	            (TMP_dWidth_mm / 2) - ((Z300_BufferPlate.rgtPlate[TMP_dIndexPlate].tData.rgtCap[TMP_dCap].rgtLite[TMP_dLite].dWidth_cmm / 100) / 2)
   	            + (Z300_BufferPlate.rgtPlate[TMP_dIndexPlate].tData.rgtCap[TMP_dCap].rgtLite[TMP_dLite].dBarycenter_cmm / 100);
   	        END_IF;
   
   	        //Barycenter used, with inversion (IN FC)
   
   	        IF TMP_xYWithBarycenter AND TMP_xYInversionLite THEN    //Barycenter used,  inversion
   	            Z300_Scada_Continuous.rgtPlate[TMP_dIndexPlate].rgtCap[TMP_dCap].rgtLite[TMP_dLite].dPositionY_mm :=
   	            (TMP_dWidth_mm / 2) - ((Z300_BufferPlate.rgtPlate[TMP_dIndexPlate].tData.rgtCap[TMP_dCap].rgtLite[TMP_dLite].dWidth_cmm / 100) / 2)
   	            - (Z300_BufferPlate.rgtPlate[TMP_dIndexPlate].tData.rgtCap[TMP_dCap].rgtLite[TMP_dLite].dBarycenter_cmm / 100);
   	        END_IF;
   	    ELSE
   	        COP(AUX_tHMI_Lite_NULL, Z300_Scada_Continuous.rgtPlate[TMP_dIndexPlate].rgtCap[TMP_dCap].rgtLite[TMP_dLite], 1);
   	    END_IF;
   	END_FOR;
   END_FOR;
   
END_ROUTINE
